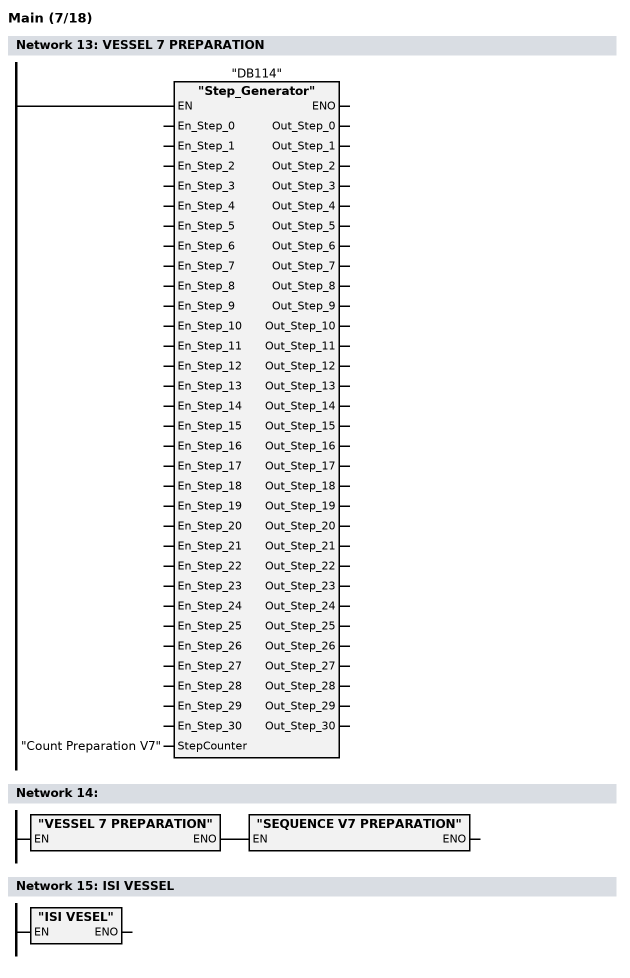
   RUNG wire#powerrail
      "DB114"(En_Step_0 :=, En_Step_1 :=, En_Step_2 :=, En_Step_3 :=, En_Step_4 :=, En_Step_5 :=, En_Step_6 :=, En_Step_7 :=, En_Step_8 :=, En_Step_9 :=, En_Step_10 :=, En_Step_11 :=, En_Step_12 :=, En_Step_13 :=, En_Step_14 :=, En_Step_15 :=, En_Step_16 :=, En_Step_17 :=, En_Step_18 :=, En_Step_19 :=, En_Step_20 :=, En_Step_21 :=, En_Step_22 :=, En_Step_23 :=, En_Step_24 :=, En_Step_25 :=, En_Step_26 :=, En_Step_27 :=, En_Step_28 :=, En_Step_29 :=, En_Step_30 :=, StepCounter := "Count Preparation V7", Out_Step_0 =>, Out_Step_1 =>, Out_Step_2 =>, Out_Step_3 =>, Out_Step_4 =>, Out_Step_5 =>, Out_Step_6 =>, Out_Step_7 =>, Out_Step_8 =>, Out_Step_9 =>, Out_Step_10 =>, Out_Step_11 =>, Out_Step_12 =>, Out_Step_13 =>, Out_Step_14 =>, Out_Step_15 =>, Out_Step_16 =>, Out_Step_17 =>, Out_Step_18 =>, Out_Step_19 =>, Out_Step_20 =>, Out_Step_21 =>, Out_Step_22 =>, Out_Step_23 =>, Out_Step_24 =>, Out_Step_25 =>, Out_Step_26 =>, Out_Step_27 =>, Out_Step_28 =>, Out_Step_29 =>, Out_Step_30 =>)
   END_RUNG
   // the same network as SCL:
   "DB114"(StepCounter := "Count Preparation V7");   // "Step_Generator"
END_REGION

REGION Network 14
   RUNG wire#powerrail
      "VESSEL 7 PREPARATION"()
      "SEQUENCE V7 PREPARATION"()
   END_RUNG
   // the same network as SCL:
   "VESSEL 7 PREPARATION"(ENO => #_w1);
   IF #_w1 THEN "SEQUENCE V7 PREPARATION"(); END_IF;
END_REGION

REGION Network 15: ISI VESSEL
   RUNG wire#powerrail
      "ISI VESEL"()
   END_RUNG
   // the same network as SCL:
   "ISI VESEL"();
END_REGION

REGION Network 16: SUPPLY
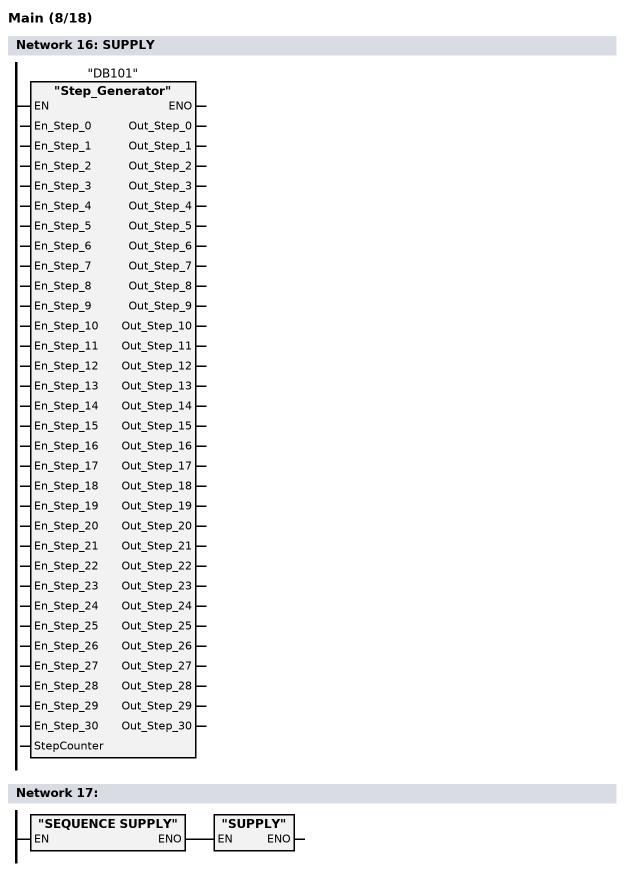
   RUNG wire#powerrail
      "DB101"(En_Step_0 :=, En_Step_1 :=, En_Step_2 :=, En_Step_3 :=, En_Step_4 :=, En_Step_5 :=, En_Step_6 :=, En_Step_7 :=, En_Step_8 :=, En_Step_9 :=, En_Step_10 :=, En_Step_11 :=, En_Step_12 :=, En_Step_13 :=, En_Step_14 :=, En_Step_15 :=, En_Step_16 :=, En_Step_17 :=, En_Step_18 :=, En_Step_19 :=, En_Step_20 :=, En_Step_21 :=, En_Step_22 :=, En_Step_23 :=, En_Step_24 :=, En_Step_25 :=, En_Step_26 :=, En_Step_27 :=, En_Step_28 :=, En_Step_29 :=, En_Step_30 :=, StepCounter :=, Out_Step_0 =>, Out_Step_1 =>, Out_Step_2 =>, Out_Step_3 =>, Out_Step_4 =>, Out_Step_5 =>, Out_Step_6 =>, Out_Step_7 =>, Out_Step_8 =>, Out_Step_9 =>, Out_Step_10 =>, Out_Step_11 =>, Out_Step_12 =>, Out_Step_13 =>, Out_Step_14 =>, Out_Step_15 =>, Out_Step_16 =>, Out_Step_17 =>, Out_Step_18 =>, Out_Step_19 =>, Out_Step_20 =>, Out_Step_21 =>, Out_Step_22 =>, Out_Step_23 =>, Out_Step_24 =>, Out_Step_25 =>, Out_Step_26 =>, Out_Step_27 =>, Out_Step_28 =>, Out_Step_29 =>, Out_Step_30 =>)
   END_RUNG
   // the same network as SCL:
   "DB101"();   // "Step_Generator"
END_REGION

REGION Network 17
   RUNG wire#powerrail
      "SEQUENCE SUPPLY"()
      "SUPPLY"()
   END_RUNG
   // the same network as SCL:
   "SEQUENCE SUPPLY"(ENO => #_w1);
   IF #_w1 THEN "SUPPLY"(); END_IF;
END_REGION

REGION Network 18: VESSEL 1
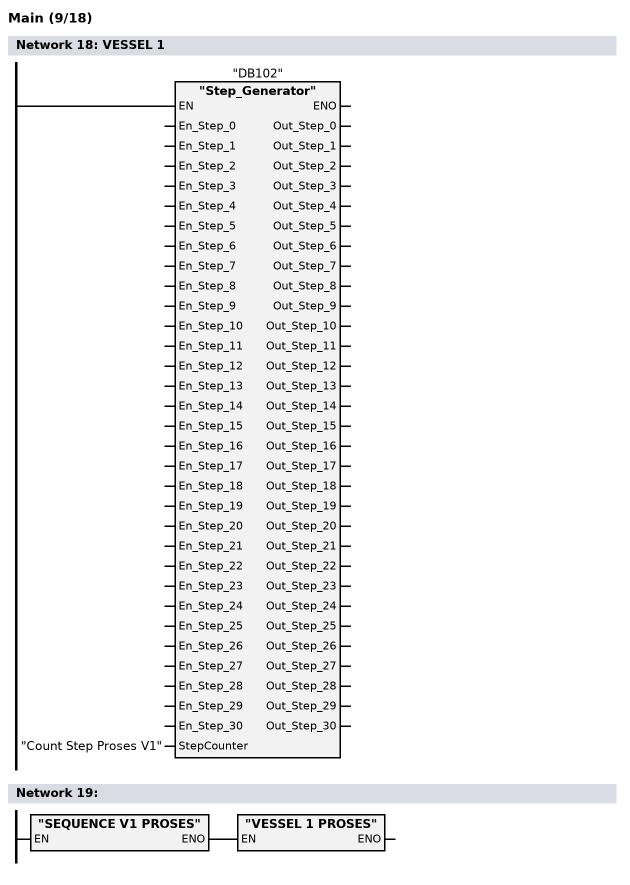
   RUNG wire#powerrail
      "DB102"(En_Step_0 :=, En_Step_1 :=, En_Step_2 :=, En_Step_3 :=, En_Step_4 :=, En_Step_5 :=, En_Step_6 :=, En_Step_7 :=, En_Step_8 :=, En_Step_9 :=, En_Step_10 :=, En_Step_11 :=, En_Step_12 :=, En_Step_13 :=, En_Step_14 :=, En_Step_15 :=, En_Step_16 :=, En_Step_17 :=, En_Step_18 :=, En_Step_19 :=, En_Step_20 :=, En_Step_21 :=, En_Step_22 :=, En_Step_23 :=, En_Step_24 :=, En_Step_25 :=, En_Step_26 :=, En_Step_27 :=, En_Step_28 :=, En_Step_29 :=, En_Step_30 :=, StepCounter := "Count Step Proses V1", Out_Step_0 =>, Out_Step_1 =>, Out_Step_2 =>, Out_Step_3 =>, Out_Step_4 =>, Out_Step_5 =>, Out_Step_6 =>, Out_Step_7 =>, Out_Step_8 =>, Out_Step_9 =>, Out_Step_10 =>, Out_Step_11 =>, Out_Step_12 =>, Out_Step_13 =>, Out_Step_14 =>, Out_Step_15 =>, Out_Step_16 =>, Out_Step_17 =>, Out_Step_18 =>, Out_Step_19 =>, Out_Step_20 =>, Out_Step_21 =>, Out_Step_22 =>, Out_Step_23 =>, Out_Step_24 =>, Out_Step_25 =>, Out_Step_26 =>, Out_Step_27 =>, Out_Step_28 =>, Out_Step_29 =>, Out_Step_30 =>)
   END_RUNG
   // the same network as SCL:
   "DB102"(StepCounter := "Count Step Proses V1");   // "Step_Generator"
END_REGION

REGION Network 19
   RUNG wire#powerrail
      "SEQUENCE V1 PROSES"()
      "VESSEL 1 PROSES"()
   END_RUNG
   // the same network as SCL:
   "SEQUENCE V1 PROSES"(ENO => #_w1);
   IF #_w1 THEN "VESSEL 1 PROSES"(); END_IF;
END_REGION

REGION Network 20: TRANSFER
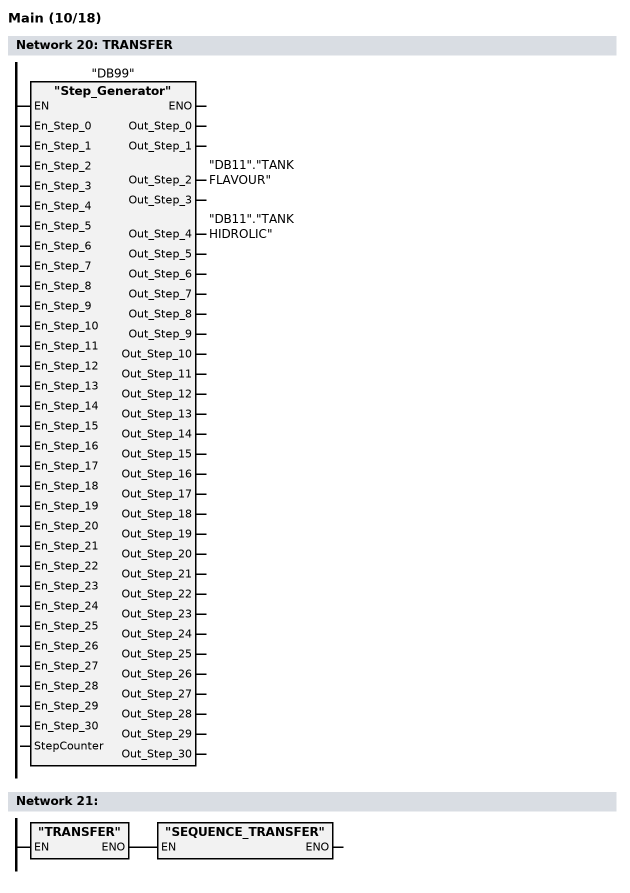
   RUNG wire#powerrail
      "DB99"(En_Step_0 :=, En_Step_1 :=, En_Step_2 :=, En_Step_3 :=, En_Step_4 :=, En_Step_5 :=, En_Step_6 :=, En_Step_7 :=, En_Step_8 :=, En_Step_9 :=, En_Step_10 :=, En_Step_11 :=, En_Step_12 :=, En_Step_13 :=, En_Step_14 :=, En_Step_15 :=, En_Step_16 :=, En_Step_17 :=, En_Step_18 :=, En_Step_19 :=, En_Step_20 :=, En_Step_21 :=, En_Step_22 :=, En_Step_23 :=, En_Step_24 :=, En_Step_25 :=, En_Step_26 :=, En_Step_27 :=, En_Step_28 :=, En_Step_29 :=, En_Step_30 :=, StepCounter :=, Out_Step_0 =>, Out_Step_1 =>, Out_Step_2 => "DB11"."TANK FLAVOUR", Out_Step_3 =>, Out_Step_4 => "DB11"."TANK HIDROLIC", Out_Step_5 =>, Out_Step_6 =>, Out_Step_7 =>, Out_Step_8 =>, Out_Step_9 =>, Out_Step_10 =>, Out_Step_11 =>, Out_Step_12 =>, Out_Step_13 =>, Out_Step_14 =>, Out_Step_15 =>, Out_Step_16 =>, Out_Step_17 =>, Out_Step_18 =>, Out_Step_19 =>, Out_Step_20 =>, Out_Step_21 =>, Out_Step_22 =>, Out_Step_23 =>, Out_Step_24 =>, Out_Step_25 =>, Out_Step_26 =>, Out_Step_27 =>, Out_Step_28 =>, Out_Step_29 =>, Out_Step_30 =>)
   END_RUNG
   // the same network as SCL:
   "DB99"(Out_Step_2 => "DB11"."TANK FLAVOUR", Out_Step_4 => "DB11"."TANK HIDROLIC");   // "Step_Generator"
END_REGION

REGION Network 21
   RUNG wire#powerrail
      "TRANSFER"()
      "SEQUENCE_TRANSFER"()
   END_RUNG
   // the same network as SCL:
   "TRANSFER"(ENO => #_w1);
   IF #_w1 THEN "SEQUENCE_TRANSFER"(); END_IF;
END_REGION

REGION Network 22: VESSEL 2
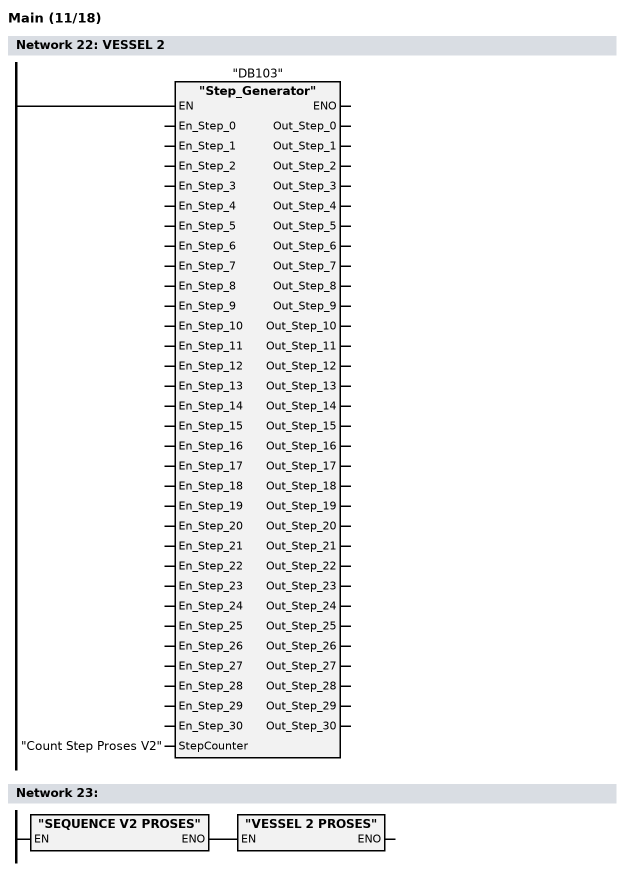
   RUNG wire#powerrail
      "DB103"(En_Step_0 :=, En_Step_1 :=, En_Step_2 :=, En_Step_3 :=, En_Step_4 :=, En_Step_5 :=, En_Step_6 :=, En_Step_7 :=, En_Step_8 :=, En_Step_9 :=, En_Step_10 :=, En_Step_11 :=, En_Step_12 :=, En_Step_13 :=, En_Step_14 :=, En_Step_15 :=, En_Step_16 :=, En_Step_17 :=, En_Step_18 :=, En_Step_19 :=, En_Step_20 :=, En_Step_21 :=, En_Step_22 :=, En_Step_23 :=, En_Step_24 :=, En_Step_25 :=, En_Step_26 :=, En_Step_27 :=, En_Step_28 :=, En_Step_29 :=, En_Step_30 :=, StepCounter := "Count Step Proses V2", Out_Step_0 =>, Out_Step_1 =>, Out_Step_2 =>, Out_Step_3 =>, Out_Step_4 =>, Out_Step_5 =>, Out_Step_6 =>, Out_Step_7 =>, Out_Step_8 =>, Out_Step_9 =>, Out_Step_10 =>, Out_Step_11 =>, Out_Step_12 =>, Out_Step_13 =>, Out_Step_14 =>, Out_Step_15 =>, Out_Step_16 =>, Out_Step_17 =>, Out_Step_18 =>, Out_Step_19 =>, Out_Step_20 =>, Out_Step_21 =>, Out_Step_22 =>, Out_Step_23 =>, Out_Step_24 =>, Out_Step_25 =>, Out_Step_26 =>, Out_Step_27 =>, Out_Step_28 =>, Out_Step_29 =>, Out_Step_30 =>)
   END_RUNG
   // the same network as SCL:
   "DB103"(StepCounter := "Count Step Proses V2");   // "Step_Generator"
END_REGION

REGION Network 23
   RUNG wire#powerrail
      "SEQUENCE V2 PROSES"()
      "VESSEL 2 PROSES"()
   END_RUNG
   // the same network as SCL:
   "SEQUENCE V2 PROSES"(ENO => #_w1);
   IF #_w1 THEN "VESSEL 2 PROSES"(); END_IF;
END_REGION

REGION Network 24: VESSEL 3 PROSES
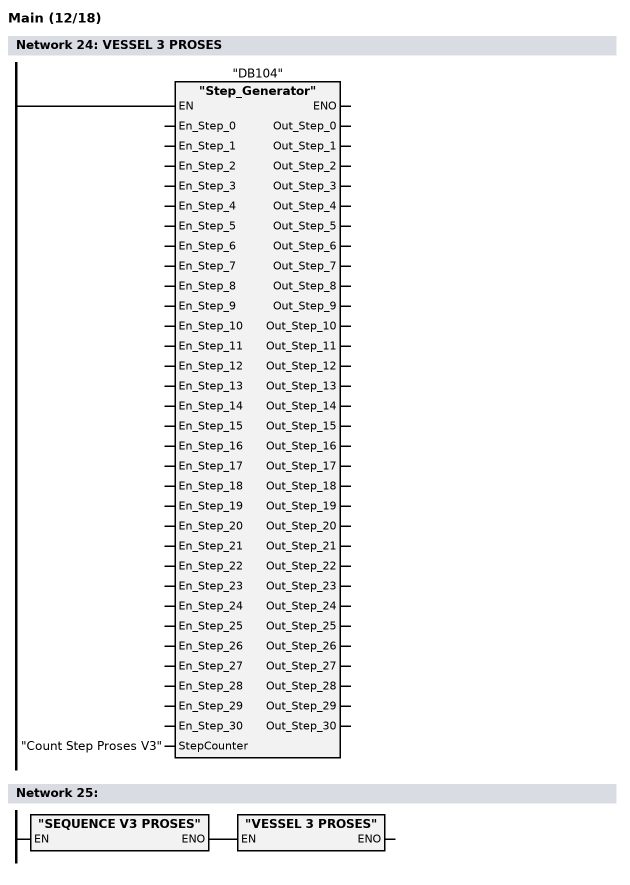
   RUNG wire#powerrail
      "DB104"(En_Step_0 :=, En_Step_1 :=, En_Step_2 :=, En_Step_3 :=, En_Step_4 :=, En_Step_5 :=, En_Step_6 :=, En_Step_7 :=, En_Step_8 :=, En_Step_9 :=, En_Step_10 :=, En_Step_11 :=, En_Step_12 :=, En_Step_13 :=, En_Step_14 :=, En_Step_15 :=, En_Step_16 :=, En_Step_17 :=, En_Step_18 :=, En_Step_19 :=, En_Step_20 :=, En_Step_21 :=, En_Step_22 :=, En_Step_23 :=, En_Step_24 :=, En_Step_25 :=, En_Step_26 :=, En_Step_27 :=, En_Step_28 :=, En_Step_29 :=, En_Step_30 :=, StepCounter := "Count Step Proses V3", Out_Step_0 =>, Out_Step_1 =>, Out_Step_2 =>, Out_Step_3 =>, Out_Step_4 =>, Out_Step_5 =>, Out_Step_6 =>, Out_Step_7 =>, Out_Step_8 =>, Out_Step_9 =>, Out_Step_10 =>, Out_Step_11 =>, Out_Step_12 =>, Out_Step_13 =>, Out_Step_14 =>, Out_Step_15 =>, Out_Step_16 =>, Out_Step_17 =>, Out_Step_18 =>, Out_Step_19 =>, Out_Step_20 =>, Out_Step_21 =>, Out_Step_22 =>, Out_Step_23 =>, Out_Step_24 =>, Out_Step_25 =>, Out_Step_26 =>, Out_Step_27 =>, Out_Step_28 =>, Out_Step_29 =>, Out_Step_30 =>)
   END_RUNG
   // the same network as SCL:
   "DB104"(StepCounter := "Count Step Proses V3");   // "Step_Generator"
END_REGION

REGION Network 25
   RUNG wire#powerrail
      "SEQUENCE V3 PROSES"()
      "VESSEL 3 PROSES"()
   END_RUNG
   // the same network as SCL:
   "SEQUENCE V3 PROSES"(ENO => #_w1);
   IF #_w1 THEN "VESSEL 3 PROSES"(); END_IF;
END_REGION

REGION Network 26: VESSEL 4
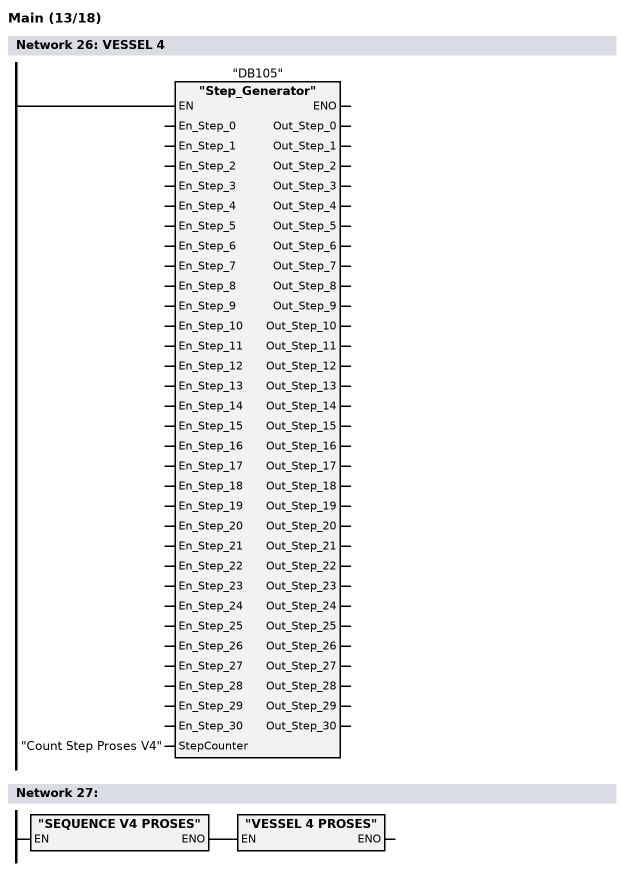
   RUNG wire#powerrail
      "DB105"(En_Step_0 :=, En_Step_1 :=, En_Step_2 :=, En_Step_3 :=, En_Step_4 :=, En_Step_5 :=, En_Step_6 :=, En_Step_7 :=, En_Step_8 :=, En_Step_9 :=, En_Step_10 :=, En_Step_11 :=, En_Step_12 :=, En_Step_13 :=, En_Step_14 :=, En_Step_15 :=, En_Step_16 :=, En_Step_17 :=, En_Step_18 :=, En_Step_19 :=, En_Step_20 :=, En_Step_21 :=, En_Step_22 :=, En_Step_23 :=, En_Step_24 :=, En_Step_25 :=, En_Step_26 :=, En_Step_27 :=, En_Step_28 :=, En_Step_29 :=, En_Step_30 :=, StepCounter := "Count Step Proses V4", Out_Step_0 =>, Out_Step_1 =>, Out_Step_2 =>, Out_Step_3 =>, Out_Step_4 =>, Out_Step_5 =>, Out_Step_6 =>, Out_Step_7 =>, Out_Step_8 =>, Out_Step_9 =>, Out_Step_10 =>, Out_Step_11 =>, Out_Step_12 =>, Out_Step_13 =>, Out_Step_14 =>, Out_Step_15 =>, Out_Step_16 =>, Out_Step_17 =>, Out_Step_18 =>, Out_Step_19 =>, Out_Step_20 =>, Out_Step_21 =>, Out_Step_22 =>, Out_Step_23 =>, Out_Step_24 =>, Out_Step_25 =>, Out_Step_26 =>, Out_Step_27 =>, Out_Step_28 =>, Out_Step_29 =>, Out_Step_30 =>)
   END_RUNG
   // the same network as SCL:
   "DB105"(StepCounter := "Count Step Proses V4");   // "Step_Generator"
END_REGION

REGION Network 27
   RUNG wire#powerrail
      "SEQUENCE V4 PROSES"()
      "VESSEL 4 PROSES"()
   END_RUNG
   // the same network as SCL:
   "SEQUENCE V4 PROSES"(ENO => #_w1);
   IF #_w1 THEN "VESSEL 4 PROSES"(); END_IF;
END_REGION

REGION Network 28: VESSEL 5
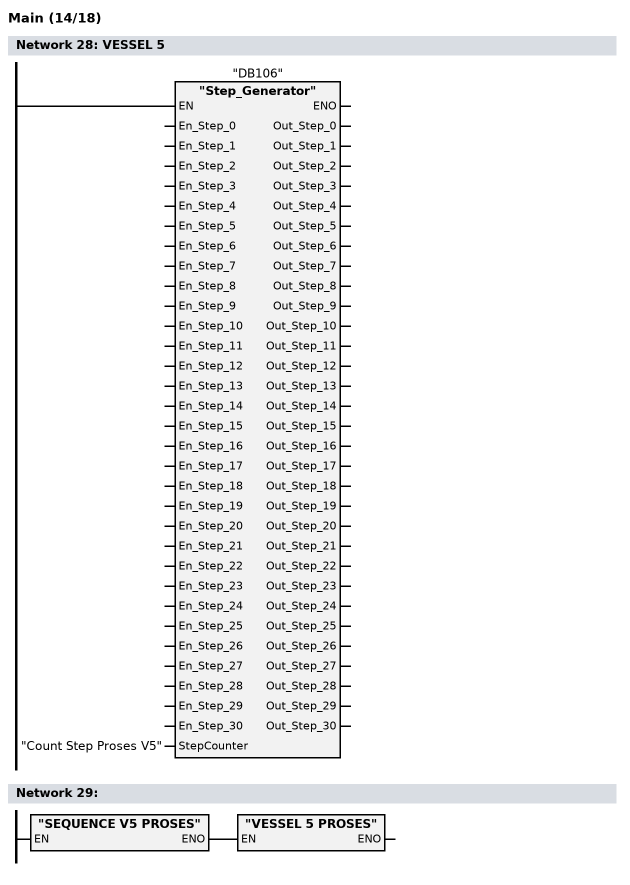
   RUNG wire#powerrail
      "DB106"(En_Step_0 :=, En_Step_1 :=, En_Step_2 :=, En_Step_3 :=, En_Step_4 :=, En_Step_5 :=, En_Step_6 :=, En_Step_7 :=, En_Step_8 :=, En_Step_9 :=, En_Step_10 :=, En_Step_11 :=, En_Step_12 :=, En_Step_13 :=, En_Step_14 :=, En_Step_15 :=, En_Step_16 :=, En_Step_17 :=, En_Step_18 :=, En_Step_19 :=, En_Step_20 :=, En_Step_21 :=, En_Step_22 :=, En_Step_23 :=, En_Step_24 :=, En_Step_25 :=, En_Step_26 :=, En_Step_27 :=, En_Step_28 :=, En_Step_29 :=, En_Step_30 :=, StepCounter := "Count Step Proses V5", Out_Step_0 =>, Out_Step_1 =>, Out_Step_2 =>, Out_Step_3 =>, Out_Step_4 =>, Out_Step_5 =>, Out_Step_6 =>, Out_Step_7 =>, Out_Step_8 =>, Out_Step_9 =>, Out_Step_10 =>, Out_Step_11 =>, Out_Step_12 =>, Out_Step_13 =>, Out_Step_14 =>, Out_Step_15 =>, Out_Step_16 =>, Out_Step_17 =>, Out_Step_18 =>, Out_Step_19 =>, Out_Step_20 =>, Out_Step_21 =>, Out_Step_22 =>, Out_Step_23 =>, Out_Step_24 =>, Out_Step_25 =>, Out_Step_26 =>, Out_Step_27 =>, Out_Step_28 =>, Out_Step_29 =>, Out_Step_30 =>)
   END_RUNG
   // the same network as SCL:
   "DB106"(StepCounter := "Count Step Proses V5");   // "Step_Generator"
END_REGION

REGION Network 29
   RUNG wire#powerrail
      "SEQUENCE V5 PROSES"()
      "VESSEL 5 PROSES"()
   END_RUNG
   // the same network as SCL:
   "SEQUENCE V5 PROSES"(ENO => #_w1);
   IF #_w1 THEN "VESSEL 5 PROSES"(); END_IF;
END_REGION

REGION Network 30: VESSEL 6
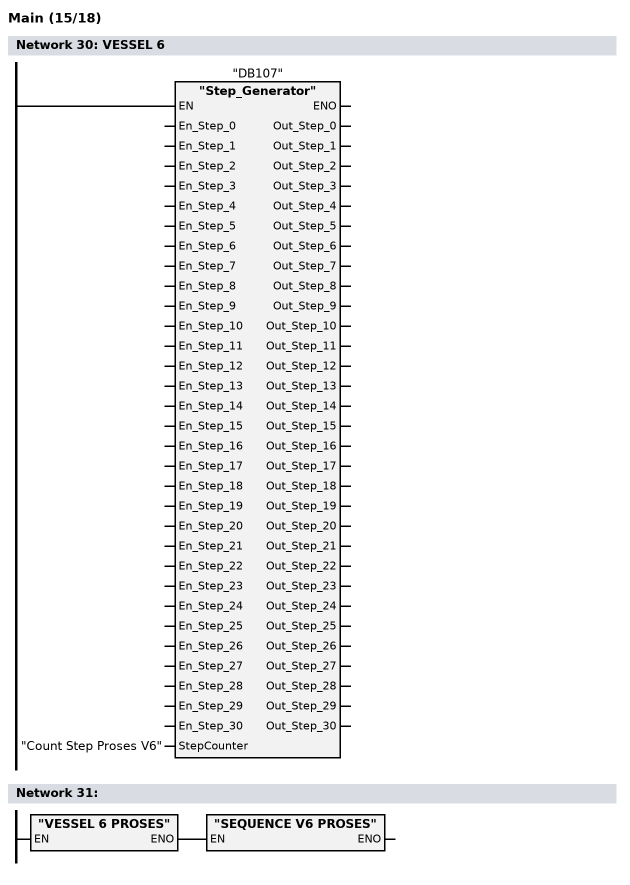
   RUNG wire#powerrail
      "DB107"(En_Step_0 :=, En_Step_1 :=, En_Step_2 :=, En_Step_3 :=, En_Step_4 :=, En_Step_5 :=, En_Step_6 :=, En_Step_7 :=, En_Step_8 :=, En_Step_9 :=, En_Step_10 :=, En_Step_11 :=, En_Step_12 :=, En_Step_13 :=, En_Step_14 :=, En_Step_15 :=, En_Step_16 :=, En_Step_17 :=, En_Step_18 :=, En_Step_19 :=, En_Step_20 :=, En_Step_21 :=, En_Step_22 :=, En_Step_23 :=, En_Step_24 :=, En_Step_25 :=, En_Step_26 :=, En_Step_27 :=, En_Step_28 :=, En_Step_29 :=, En_Step_30 :=, StepCounter := "Count Step Proses V6", Out_Step_0 =>, Out_Step_1 =>, Out_Step_2 =>, Out_Step_3 =>, Out_Step_4 =>, Out_Step_5 =>, Out_Step_6 =>, Out_Step_7 =>, Out_Step_8 =>, Out_Step_9 =>, Out_Step_10 =>, Out_Step_11 =>, Out_Step_12 =>, Out_Step_13 =>, Out_Step_14 =>, Out_Step_15 =>, Out_Step_16 =>, Out_Step_17 =>, Out_Step_18 =>, Out_Step_19 =>, Out_Step_20 =>, Out_Step_21 =>, Out_Step_22 =>, Out_Step_23 =>, Out_Step_24 =>, Out_Step_25 =>, Out_Step_26 =>, Out_Step_27 =>, Out_Step_28 =>, Out_Step_29 =>, Out_Step_30 =>)
   END_RUNG
   // the same network as SCL:
   "DB107"(StepCounter := "Count Step Proses V6");   // "Step_Generator"
END_REGION

REGION Network 31
   RUNG wire#powerrail
      "VESSEL 6 PROSES"()
      "SEQUENCE V6 PROSES"()
   END_RUNG
   // the same network as SCL:
   "VESSEL 6 PROSES"(ENO => #_w1);
   IF #_w1 THEN "SEQUENCE V6 PROSES"(); END_IF;
END_REGION

REGION Network 32: VESSEL 7
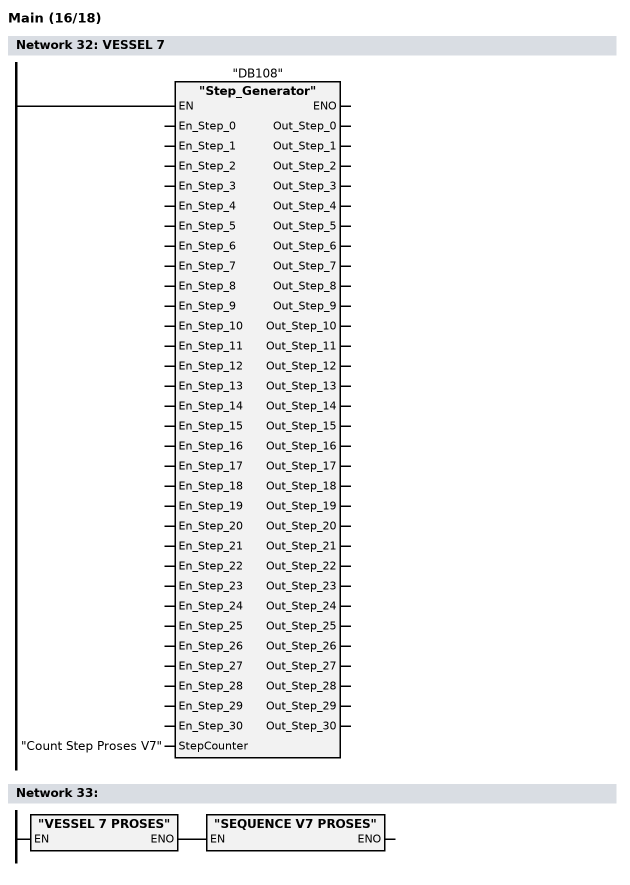
   RUNG wire#powerrail
      "DB108"(En_Step_0 :=, En_Step_1 :=, En_Step_2 :=, En_Step_3 :=, En_Step_4 :=, En_Step_5 :=, En_Step_6 :=, En_Step_7 :=, En_Step_8 :=, En_Step_9 :=, En_Step_10 :=, En_Step_11 :=, En_Step_12 :=, En_Step_13 :=, En_Step_14 :=, En_Step_15 :=, En_Step_16 :=, En_Step_17 :=, En_Step_18 :=, En_Step_19 :=, En_Step_20 :=, En_Step_21 :=, En_Step_22 :=, En_Step_23 :=, En_Step_24 :=, En_Step_25 :=, En_Step_26 :=, En_Step_27 :=, En_Step_28 :=, En_Step_29 :=, En_Step_30 :=, StepCounter := "Count Step Proses V7", Out_Step_0 =>, Out_Step_1 =>, Out_Step_2 =>, Out_Step_3 =>, Out_Step_4 =>, Out_Step_5 =>, Out_Step_6 =>, Out_Step_7 =>, Out_Step_8 =>, Out_Step_9 =>, Out_Step_10 =>, Out_Step_11 =>, Out_Step_12 =>, Out_Step_13 =>, Out_Step_14 =>, Out_Step_15 =>, Out_Step_16 =>, Out_Step_17 =>, Out_Step_18 =>, Out_Step_19 =>, Out_Step_20 =>, Out_Step_21 =>, Out_Step_22 =>, Out_Step_23 =>, Out_Step_24 =>, Out_Step_25 =>, Out_Step_26 =>, Out_Step_27 =>, Out_Step_28 =>, Out_Step_29 =>, Out_Step_30 =>)
   END_RUNG
   // the same network as SCL:
   "DB108"(StepCounter := "Count Step Proses V7");   // "Step_Generator"
END_REGION

REGION Network 33
   RUNG wire#powerrail
      "VESSEL 7 PROSES"()
      "SEQUENCE V7 PROSES"()
   END_RUNG
   // the same network as SCL:
   "VESSEL 7 PROSES"(ENO => #_w1);
   IF #_w1 THEN "SEQUENCE V7 PROSES"(); END_IF;
END_REGION

REGION Network 34: CLEAN
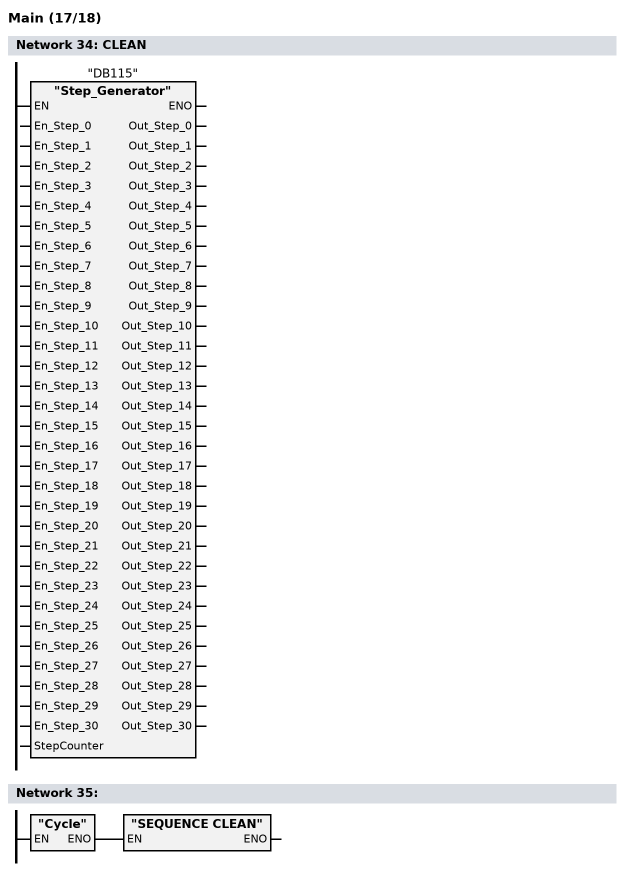
   RUNG wire#powerrail
      "DB115"(En_Step_0 :=, En_Step_1 :=, En_Step_2 :=, En_Step_3 :=, En_Step_4 :=, En_Step_5 :=, En_Step_6 :=, En_Step_7 :=, En_Step_8 :=, En_Step_9 :=, En_Step_10 :=, En_Step_11 :=, En_Step_12 :=, En_Step_13 :=, En_Step_14 :=, En_Step_15 :=, En_Step_16 :=, En_Step_17 :=, En_Step_18 :=, En_Step_19 :=, En_Step_20 :=, En_Step_21 :=, En_Step_22 :=, En_Step_23 :=, En_Step_24 :=, En_Step_25 :=, En_Step_26 :=, En_Step_27 :=, En_Step_28 :=, En_Step_29 :=, En_Step_30 :=, StepCounter :=, Out_Step_0 =>, Out_Step_1 =>, Out_Step_2 =>, Out_Step_3 =>, Out_Step_4 =>, Out_Step_5 =>, Out_Step_6 =>, Out_Step_7 =>, Out_Step_8 =>, Out_Step_9 =>, Out_Step_10 =>, Out_Step_11 =>, Out_Step_12 =>, Out_Step_13 =>, Out_Step_14 =>, Out_Step_15 =>, Out_Step_16 =>, Out_Step_17 =>, Out_Step_18 =>, Out_Step_19 =>, Out_Step_20 =>, Out_Step_21 =>, Out_Step_22 =>, Out_Step_23 =>, Out_Step_24 =>, Out_Step_25 =>, Out_Step_26 =>, Out_Step_27 =>, Out_Step_28 =>, Out_Step_29 =>, Out_Step_30 =>)
   END_RUNG
   // the same network as SCL:
   "DB115"();   // "Step_Generator"
END_REGION

REGION Network 35
   RUNG wire#powerrail
      "Cycle"()
      "SEQUENCE CLEAN"()
   END_RUNG
   // the same network as SCL:
   "Cycle"(ENO => #_w1);
   IF #_w1 THEN "SEQUENCE CLEAN"(); END_IF;
END_REGION

REGION Network 36
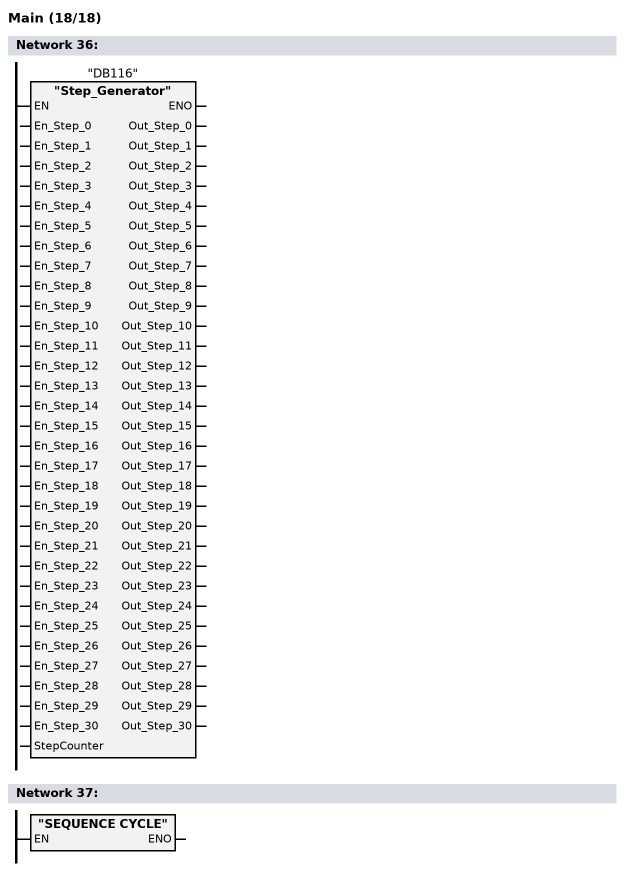
   RUNG wire#powerrail
      "DB116"(En_Step_0 :=, En_Step_1 :=, En_Step_2 :=, En_Step_3 :=, En_Step_4 :=, En_Step_5 :=, En_Step_6 :=, En_Step_7 :=, En_Step_8 :=, En_Step_9 :=, En_Step_10 :=, En_Step_11 :=, En_Step_12 :=, En_Step_13 :=, En_Step_14 :=, En_Step_15 :=, En_Step_16 :=, En_Step_17 :=, En_Step_18 :=, En_Step_19 :=, En_Step_20 :=, En_Step_21 :=, En_Step_22 :=, En_Step_23 :=, En_Step_24 :=, En_Step_25 :=, En_Step_26 :=, En_Step_27 :=, En_Step_28 :=, En_Step_29 :=, En_Step_30 :=, StepCounter :=, Out_Step_0 =>, Out_Step_1 =>, Out_Step_2 =>, Out_Step_3 =>, Out_Step_4 =>, Out_Step_5 =>, Out_Step_6 =>, Out_Step_7 =>, Out_Step_8 =>, Out_Step_9 =>, Out_Step_10 =>, Out_Step_11 =>, Out_Step_12 =>, Out_Step_13 =>, Out_Step_14 =>, Out_Step_15 =>, Out_Step_16 =>, Out_Step_17 =>, Out_Step_18 =>, Out_Step_19 =>, Out_Step_20 =>, Out_Step_21 =>, Out_Step_22 =>, Out_Step_23 =>, Out_Step_24 =>, Out_Step_25 =>, Out_Step_26 =>, Out_Step_27 =>, Out_Step_28 =>, Out_Step_29 =>, Out_Step_30 =>)
   END_RUNG
   // the same network as SCL:
   "DB116"();   // "Step_Generator"
END_REGION

REGION Network 37
   RUNG wire#powerrail
      "SEQUENCE CYCLE"()
   END_RUNG
   // the same network as SCL:
   "SEQUENCE CYCLE"();
END_REGION
END_ORGANIZATION_BLOCK

(* ===== HMI "HMI_RT_1" =====
system functions are stored by id; their names below are inferred from use
connection "Connection_1": ETHERNET, S7_1500_OMS
connection "HMI_Connection_1": ETHERNET, S7_1500_OMS

HMI tags "Default tag table"
   "testag" : Bool, internal
   "preparation" : Bool AT %M100.0, 1 s
   "pressure vessel 1" : Int AT %MW200, 1 s
   "pressure vessel 2" : Int AT %MW202, 1 s
   "pressure vessel 3" : Int AT %MW204, 1 s
   "pressure vessel 4" : Int AT %MW206, 1 s
   "pressure vessel 5" : Int AT %MW208, 1 s
   "pressure vessel 6" : Int AT %MW210, 1 s
   "pressure vessel 7" : Int AT %MW212, 1 s
   "reset" : Bool AT %M100.5, 1 s
   "PROSES" : Bool AT %M100.4, 1 s
   "RESET 2" : Bool AT %M100.6, 1 s
   "pressure steam supply" : Int AT %MW230, 1 s
   "temperature THE 1" : Int AT %MW164, 1 s
   "temperature THE 2" : Int AT %MW166, 1 s
   "temperature vesel 1" : Int AT %MW240, 1 s
   "temperature vesel 2" : Int AT %MW242, 1 s
   "temperature vesel 3" : Int AT %MW244, 1 s
   "temperature vesel 4" : Int AT %MW246, 1 s
   "temperature vesel 5" : Int AT %MW248, 1 s
   "temperature vesel 6" : Int AT %MW250, 1 s
   "temperature vesel 7" : Int AT %MW252, 1 s
   "tank flavour OK" : Bool AT %DB11.DBX0.2, 1 s
   "tank hidrolic OK" : Bool AT %DB11.DBX0.3, 1 s
   "transfer" : Bool AT %M100.5, 1 s
   "PROSES_2" : Bool AT %M100.6, 1 s
   "preparation_v1" : Bool AT %M100.0, 1 s
   "preparation_v2" : Bool AT %M101.3, 1 s
   "preparation_v3" : Bool AT %M101.4, 1 s
   "preparation_v4" : Bool AT %M101.5, 1 s
   "preparation_v5" : Bool AT %M101.6, 1 s
   "preparation_v6" : Bool AT %M101.7, 1 s
   "preparation_v7" : Bool AT %M102.0, 1 s
   "proses_v1" : Bool AT %M100.4, 1 s
   "proses_v2" : Bool AT %M100.6, 1 s
   "proses_v3" : Bool AT %M100.7, 1 s
   "proses_v4" : Bool AT %M101.0, 1 s
   "proses_v5" : Bool AT %M101.1, 1 s
   "proses_v6" : Bool AT %M101.2, 1 s
   "proses_v7" : Bool AT %M102.7, 1 s
   "cyclecounter" : Int AT %DB11.DBW2, 1 s
   "mode" : Bool AT %DB11.DBX4.7, 1 s
   "reset_cycle" : Bool AT %M103.0, 1 s
   "supply" : Bool AT %M100.3, 1 s
   "isi_vesel_start" : Bool AT %M100.2, 1 s
   "Count Step Proses V1" : Int = PLC "Count Step Proses V1" AT %MW140, 1 s
   "EMERGENCY" : Bool AT %M103.1, 1 s
